   4659: 'Spare_Fault_4659', class No Acknowledgement, trigger "DB302_HMI_Faults_Carrier72_Faults_3" bit 2
   4660: 'Spare_Fault_4660', class No Acknowledgement, trigger "DB302_HMI_Faults_Carrier72_Faults_3" bit 3
   4661: 'Spare_Fault_4661', class No Acknowledgement, trigger "DB302_HMI_Faults_Carrier72_Faults_3" bit 4
   4662: 'Spare_Fault_4662', class No Acknowledgement, trigger "DB302_HMI_Faults_Carrier72_Faults_3" bit 5
   4663: 'Spare_Fault_4663', class No Acknowledgement, trigger "DB302_HMI_Faults_Carrier72_Faults_3" bit 6
   4664: 'Spare_Fault_4664', class No Acknowledgement, trigger "DB302_HMI_Faults_Carrier72_Faults_3" bit 7
   4665: 'Spare_Fault_4665', class No Acknowledgement, trigger "DB302_HMI_Faults_Carrier72_Faults_3" bit 8
   4666: 'Spare_Fault_4666', class No Acknowledgement, trigger "DB302_HMI_Faults_Carrier72_Faults_3" bit 9
   4667: 'Spare_Fault_4667', class No Acknowledgement, trigger "DB302_HMI_Faults_Carrier72_Faults_3" bit 10
   4668: 'Spare_Fault_4668', class No Acknowledgement, trigger "DB302_HMI_Faults_Carrier72_Faults_3" bit 11
   4669: 'Spare_Fault_4669', class No Acknowledgement, trigger "DB302_HMI_Faults_Carrier72_Faults_3" bit 12
   4670: 'Spare_Fault_4670', class No Acknowledgement, trigger "DB302_HMI_Faults_Carrier72_Faults_3" bit 13
   4671: 'Spare_Fault_4671', class No Acknowledgement, trigger "DB302_HMI_Faults_Carrier72_Faults_3" bit 14
   4672: 'Spare_Fault_4672', class No Acknowledgement, trigger "DB302_HMI_Faults_Carrier72_Faults_3" bit 15
   4673: 'Carrier 73 Disconnect Open Power Fault DI11.0', class No Acknowledgement, trigger "DB302_HMI_Faults_Carrier73_Faults_0" bit 0
   4674: 'Carrier 73 Drive Profinet Comm Fault', class No Acknowledgement, trigger "DB302_HMI_Faults_Carrier73_Faults_0" bit 1
   4675: 'Carrier 73 Production Stop Not Reset', class No Acknowledgement, trigger "DB302_HMI_Faults_Carrier73_Faults_0" bit 2
   4676: 'Carrier 73 CB02122 Tripped', class No Acknowledgement, trigger "DB302_HMI_Faults_Carrier73_Faults_0" bit 3
   4677: 'Carrier 73 CB02123 Tripped', class No Acknowledgement, trigger "DB302_HMI_Faults_Carrier73_Faults_0" bit 4
   4678: 'Carrier 73 AUX1 CB Tripped', class No Acknowledgement, trigger "DB302_HMI_Faults_Carrier73_Faults_0" bit 5
   4679: 'Carrier 73 AUX2 CB Tripped', class No Acknowledgement, trigger "DB302_HMI_Faults_Carrier73_Faults_0" bit 6
   4680: 'Carrier 73 PLC Not Communicating', class No Acknowledgement, trigger "DB302_HMI_Faults_Carrier73_Faults_0" bit 7
   4681: 'Carrier 73 Safe Input Card Fault', class No Acknowledgement, trigger "DB302_HMI_Faults_Carrier73_Faults_0" bit 8
   4682: 'Carrier 73 Safe Output Card Fault', class No Acknowledgement, trigger "DB302_HMI_Faults_Carrier73_Faults_0" bit 9
   4683: 'Carrier 73 Standard Input Card Fault', class No Acknowledgement, trigger "DB302_HMI_Faults_Carrier73_Faults_0" bit 10
   4684: 'Carrier 73 Standard Output Card Fault', class No Acknowledgement, trigger "DB302_HMI_Faults_Carrier73_Faults_0" bit 11
   4685: 'Carrier 73 Encoder Position Fault', class No Acknowledgement, trigger "DB302_HMI_Faults_Carrier73_Faults_0" bit 12
   4686: 'Carrier 73 Encoder Internal Error', class No Acknowledgement, trigger "DB302_HMI_Faults_Carrier73_Faults_0" bit 13
   4687: 'Carrier 73 Encoder Comm Fault', class No Acknowledgement, trigger "DB302_HMI_Faults_Carrier73_Faults_0" bit 14
   4688: 'Carrier 73 HMI Comm Fault', class No Acknowledgement, trigger "DB302_HMI_Faults_Carrier73_Faults_0" bit 15
   4689: 'Carrier 73 Crash Detection Fault', class No Acknowledgement, trigger "DB302_HMI_Faults_Carrier73_Faults_1" bit 0
   4690: 'Carrier 73 Carrier Number Invalid', class No Acknowledgement, trigger "DB302_HMI_Faults_Carrier73_Faults_1" bit 1
   4691: 'Carrier 73 Drive: PROFINET configuration error', class No Acknowledgement, trigger "DB302_HMI_Faults_Carrier73_Faults_1" bit 2
   4692: 'Carrier 73 Drive: Error internal communications', class No Acknowledgement, trigger "DB302_HMI_Faults_Carrier73_Faults_1" bit 3
   4693: 'Carrier 73 Drive: Motor overtemperature', class No Acknowledgement, trigger "DB302_HMI_Faults_Carrier73_Faults_1" bit 4
   4694: 'Carrier 73 Drive: Motor overcurrent', class No Acknowledgement, trigger "DB302_HMI_Faults_Carrier73_Faults_1" bit 5
   4695: 'Carrier 73 Drive: Infeed or power unit not ready', class No Acknowledgement, trigger "DB302_HMI_Faults_Carrier73_Faults_1" bit 6
   4696: 'Carrier 73 Drive: Short-circuit/ground fault detected', class No Acknowledgement, trigger "DB302_HMI_Faults_Carrier73_Faults_1" bit 7
   4697: 'Carrier 73 Drive: PROFINET Setpoint timeout', class No Acknowledgement, trigger "DB302_HMI_Faults_Carrier73_Faults_1" bit 8
   4698: 'Carrier 73 Power unit: Overcurrent', class No Acknowledgement, trigger "DB302_HMI_Faults_Carrier73_Faults_1" bit 9
   4699: 'Carrier 73 Power unit: DC link voltage overvoltage', class No Acknowledgement, trigger "DB302_HMI_Faults_Carrier73_Faults_1" bit 10
   4700: 'Carrier 73 Power unit: DC link voltage undervoltage', class No Acknowledgement, trigger "DB302_HMI_Faults_Carrier73_Faults_1" bit 11
   4701: 'Carrier 73 Power unit: Line phase failure in main circuit', class No Acknowledgement, trigger "DB302_HMI_Faults_Carrier73_Faults_1" bit 12
   4702: 'Carrier 73 Power unit: Phase failure motor cable', class No Acknowledgement, trigger "DB302_HMI_Faults_Carrier73_Faults_1" bit 13
   4703: 'Carrier 73 Power unit: Ground fault', class No Acknowledgement, trigger "DB302_HMI_Faults_Carrier73_Faults_1" bit 14
   4704: 'Spare_Fault_4704', class No Acknowledgement, trigger "DB302_HMI_Faults_Carrier73_Faults_1" bit 15
   4705: 'Carrier 73 Motion Off Fault', class No Acknowledgement, trigger "DB302_HMI_Faults_Carrier73_Faults_2" bit 0
   4706: 'Carrier 73 Motion On Fault', class No Acknowledgement, trigger "DB302_HMI_Faults_Carrier73_Faults_2" bit 1
   4707: 'Carrier 73 Spacing Fault', class No Acknowledgement, trigger "DB302_HMI_Faults_Carrier73_Faults_2" bit 2
   4708: 'Carrier 73 Duplicate Carrier Number Fault', class No Acknowledgement, trigger "DB302_HMI_Faults_Carrier73_Faults_2" bit 3
   4709: 'Spare_Fault_4709', class No Acknowledgement, trigger "DB302_HMI_Faults_Carrier73_Faults_2" bit 4
   4710: 'Spare_Fault_4710', class No Acknowledgement, trigger "DB302_HMI_Faults_Carrier73_Faults_2" bit 5
   4711: 'Spare_Fault_4711', class No Acknowledgement, trigger "DB302_HMI_Faults_Carrier73_Faults_2" bit 6
   4712: 'Spare_Fault_4712', class No Acknowledgement, trigger "DB302_HMI_Faults_Carrier73_Faults_2" bit 7
   4713: 'Spare_Fault_4713', class No Acknowledgement, trigger "DB302_HMI_Faults_Carrier73_Faults_2" bit 8
   4714: 'Spare_Fault_4714', class No Acknowledgement, trigger "DB302_HMI_Faults_Carrier73_Faults_2" bit 9
   4715: 'Spare_Fault_4715', class No Acknowledgement, trigger "DB302_HMI_Faults_Carrier73_Faults_2" bit 10
   4716: 'Spare_Fault_4716', class No Acknowledgement, trigger "DB302_HMI_Faults_Carrier73_Faults_2" bit 11
   4717: 'Spare_Fault_4717', class No Acknowledgement, trigger "DB302_HMI_Faults_Carrier73_Faults_2" bit 12
   4718: 'Spare_Fault_4718', class No Acknowledgement, trigger "DB302_HMI_Faults_Carrier73_Faults_2" bit 13
   4719: 'Spare_Fault_4719', class No Acknowledgement, trigger "DB302_HMI_Faults_Carrier73_Faults_2" bit 14
   4720: 'Spare_Fault_4720', class No Acknowledgement, trigger "DB302_HMI_Faults_Carrier73_Faults_2" bit 15
   4721: 'Spare_Fault_4721', class No Acknowledgement, trigger "DB302_HMI_Faults_Carrier73_Faults_3" bit 0
   4722: 'Spare_Fault_4722', class No Acknowledgement, trigger "DB302_HMI_Faults_Carrier73_Faults_3" bit 1
   4723: 'Spare_Fault_4723', class No Acknowledgement, trigger "DB302_HMI_Faults_Carrier73_Faults_3" bit 2
   4724: 'Spare_Fault_4724', class No Acknowledgement, trigger "DB302_HMI_Faults_Carrier73_Faults_3" bit 3
   4725: 'Spare_Fault_4725', class No Acknowledgement, trigger "DB302_HMI_Faults_Carrier73_Faults_3" bit 4
   4726: 'Spare_Fault_4726', class No Acknowledgement, trigger "DB302_HMI_Faults_Carrier73_Faults_3" bit 5
   4727: 'Spare_Fault_4727', class No Acknowledgement, trigger "DB302_HMI_Faults_Carrier73_Faults_3" bit 6
   4728: 'Spare_Fault_4728', class No Acknowledgement, trigger "DB302_HMI_Faults_Carrier73_Faults_3" bit 7
   4729: 'Spare_Fault_4729', class No Acknowledgement, trigger "DB302_HMI_Faults_Carrier73_Faults_3" bit 8
   4730: 'Spare_Fault_4730', class No Acknowledgement, trigger "DB302_HMI_Faults_Carrier73_Faults_3" bit 9
   4731: 'Spare_Fault_4731', class No Acknowledgement, trigger "DB302_HMI_Faults_Carrier73_Faults_3" bit 10
   4732: 'Spare_Fault_4732', class No Acknowledgement, trigger "DB302_HMI_Faults_Carrier73_Faults_3" bit 11
   4733: 'Spare_Fault_4733', class No Acknowledgement, trigger "DB302_HMI_Faults_Carrier73_Faults_3" bit 12
   4734: 'Spare_Fault_4734', class No Acknowledgement, trigger "DB302_HMI_Faults_Carrier73_Faults_3" bit 13
   4735: 'Spare_Fault_4735', class No Acknowledgement, trigger "DB302_HMI_Faults_Carrier73_Faults_3" bit 14
   4736: 'Spare_Fault_4736', class No Acknowledgement, trigger "DB302_HMI_Faults_Carrier73_Faults_3" bit 15
   4737: 'Carrier 74 Disconnect Open Power Fault DI11.0', class No Acknowledgement, trigger "DB302_HMI_Faults_Carrier74_Faults_0" bit 0
   4738: 'Carrier 74 Drive Profinet Comm Fault', class No Acknowledgement, trigger "DB302_HMI_Faults_Carrier74_Faults_0" bit 1
   4739: 'Carrier 74 Production Stop Not Reset', class No Acknowledgement, trigger "DB302_HMI_Faults_Carrier74_Faults_0" bit 2
   4740: 'Carrier 74 CB02122 Tripped', class No Acknowledgement, trigger "DB302_HMI_Faults_Carrier74_Faults_0" bit 3
   4741: 'Carrier 74 CB02123 Tripped', class No Acknowledgement, trigger "DB302_HMI_Faults_Carrier74_Faults_0" bit 4
   4742: 'Carrier 74 AUX1 CB Tripped', class No Acknowledgement, trigger "DB302_HMI_Faults_Carrier74_Faults_0" bit 5
   4743: 'Carrier 74 AUX2 CB Tripped', class No Acknowledgement, trigger "DB302_HMI_Faults_Carrier74_Faults_0" bit 6
   4744: 'Carrier 74 PLC Not Communicating', class No Acknowledgement, trigger "DB302_HMI_Faults_Carrier74_Faults_0" bit 7
   4745: 'Carrier 74 Safe Input Card Fault', class No Acknowledgement, trigger "DB302_HMI_Faults_Carrier74_Faults_0" bit 8
   4746: 'Carrier 74 Safe Output Card Fault', class No Acknowledgement, trigger "DB302_HMI_Faults_Carrier74_Faults_0" bit 9
   4747: 'Carrier 74 Standard Input Card Fault', class No Acknowledgement, trigger "DB302_HMI_Faults_Carrier74_Faults_0" bit 10
   4748: 'Carrier 74 Standard Output Card Fault', class No Acknowledgement, trigger "DB302_HMI_Faults_Carrier74_Faults_0" bit 11
   4749: 'Carrier 74 Encoder Position Fault', class No Acknowledgement, trigger "DB302_HMI_Faults_Carrier74_Faults_0" bit 12
   4750: 'Carrier 74 Encoder Internal Error', class No Acknowledgement, trigger "DB302_HMI_Faults_Carrier74_Faults_0" bit 13
   4751: 'Carrier 74 Encoder Comm Fault', class No Acknowledgement, trigger "DB302_HMI_Faults_Carrier74_Faults_0" bit 14
   4752: 'Carrier 74 HMI Comm Fault', class No Acknowledgement, trigger "DB302_HMI_Faults_Carrier74_Faults_0" bit 15
   4753: 'Carrier 74 Crash Detection Fault', class No Acknowledgement, trigger "DB302_HMI_Faults_Carrier74_Faults_1" bit 0
   4754: 'Carrier 74 Carrier Number Invalid', class No Acknowledgement, trigger "DB302_HMI_Faults_Carrier74_Faults_1" bit 1
   4755: 'Carrier 74 Drive: PROFINET configuration error', class No Acknowledgement, trigger "DB302_HMI_Faults_Carrier74_Faults_1" bit 2
   4756: 'Carrier 74 Drive: Error internal communications', class No Acknowledgement, trigger "DB302_HMI_Faults_Carrier74_Faults_1" bit 3
   4757: 'Carrier 74 Drive: Motor overtemperature', class No Acknowledgement, trigger "DB302_HMI_Faults_Carrier74_Faults_1" bit 4
   4758: 'Carrier 74 Drive: Motor overcurrent', class No Acknowledgement, trigger "DB302_HMI_Faults_Carrier74_Faults_1" bit 5
   4759: 'Carrier 74 Drive: Infeed or power unit not ready', class No Acknowledgement, trigger "DB302_HMI_Faults_Carrier74_Faults_1" bit 6
   4760: 'Carrier 74 Drive: Short-circuit/ground fault detected', class No Acknowledgement, trigger "DB302_HMI_Faults_Carrier74_Faults_1" bit 7
   4761: 'Carrier 74 Drive: PROFINET Setpoint timeout', class No Acknowledgement, trigger "DB302_HMI_Faults_Carrier74_Faults_1" bit 8
   4762: 'Carrier 74 Power unit: Overcurrent', class No Acknowledgement, trigger "DB302_HMI_Faults_Carrier74_Faults_1" bit 9
   4763: 'Carrier 74 Power unit: DC link voltage overvoltage', class No Acknowledgement, trigger "DB302_HMI_Faults_Carrier74_Faults_1" bit 10
   4764: 'Carrier 74 Power unit: DC link voltage undervoltage', class No Acknowledgement, trigger "DB302_HMI_Faults_Carrier74_Faults_1" bit 11
   4765: 'Carrier 74 Power unit: Line phase failure in main circuit', class No Acknowledgement, trigger "DB302_HMI_Faults_Carrier74_Faults_1" bit 12
   4766: 'Carrier 74 Power unit: Phase failure motor cable', class No Acknowledgement, trigger "DB302_HMI_Faults_Carrier74_Faults_1" bit 13
   4767: 'Carrier 74 Power unit: Ground fault', class No Acknowledgement, trigger "DB302_HMI_Faults_Carrier74_Faults_1" bit 14
   4768: 'Spare_Fault_4768', class No Acknowledgement, trigger "DB302_HMI_Faults_Carrier74_Faults_1" bit 15
   4769: 'Carrier 74 Motion Off Fault', class No Acknowledgement, trigger "DB302_HMI_Faults_Carrier74_Faults_2" bit 0
   4770: 'Carrier 74 Motion On Fault', class No Acknowledgement, trigger "DB302_HMI_Faults_Carrier74_Faults_2" bit 1
   4771: 'Carrier 74 Spacing Fault', class No Acknowledgement, trigger "DB302_HMI_Faults_Carrier74_Faults_2" bit 2
   4772: 'Carrier 74 Duplicate Carrier Number Fault', class No Acknowledgement, trigger "DB302_HMI_Faults_Carrier74_Faults_2" bit 3
   4773: 'Spare_Fault_4773', class No Acknowledgement, trigger "DB302_HMI_Faults_Carrier74_Faults_2" bit 4
   4774: 'Spare_Fault_4774', class No Acknowledgement, trigger "DB302_HMI_Faults_Carrier74_Faults_2" bit 5
   4775: 'Spare_Fault_4775', class No Acknowledgement, trigger "DB302_HMI_Faults_Carrier74_Faults_2" bit 6
   4776: 'Spare_Fault_4776', class No Acknowledgement, trigger "DB302_HMI_Faults_Carrier74_Faults_2" bit 7
   4777: 'Spare_Fault_4777', class No Acknowledgement, trigger "DB302_HMI_Faults_Carrier74_Faults_2" bit 8
   4778: 'Spare_Fault_4778', class No Acknowledgement, trigger "DB302_HMI_Faults_Carrier74_Faults_2" bit 9
   4779: 'Spare_Fault_4779', class No Acknowledgement, trigger "DB302_HMI_Faults_Carrier74_Faults_2" bit 10
   4780: 'Spare_Fault_4780', class No Acknowledgement, trigger "DB302_HMI_Faults_Carrier74_Faults_2" bit 11
   4781: 'Spare_Fault_4781', class No Acknowledgement, trigger "DB302_HMI_Faults_Carrier74_Faults_2" bit 12
   4782: 'Spare_Fault_4782', class No Acknowledgement, trigger "DB302_HMI_Faults_Carrier74_Faults_2" bit 13
   4783: 'Spare_Fault_4783', class No Acknowledgement, trigger "DB302_HMI_Faults_Carrier74_Faults_2" bit 14
   4784: 'Spare_Fault_4784', class No Acknowledgement, trigger "DB302_HMI_Faults_Carrier74_Faults_2" bit 15
   4785: 'Spare_Fault_4785', class No Acknowledgement, trigger "DB302_HMI_Faults_Carrier74_Faults_3" bit 0
   4786: 'Spare_Fault_4786', class No Acknowledgement, trigger "DB302_HMI_Faults_Carrier74_Faults_3" bit 1
   4787: 'Spare_Fault_4787', class No Acknowledgement, trigger "DB302_HMI_Faults_Carrier74_Faults_3" bit 2
   4788: 'Spare_Fault_4788', class No Acknowledgement, trigger "DB302_HMI_Faults_Carrier74_Faults_3" bit 3
   4789: 'Spare_Fault_4789', class No Acknowledgement, trigger "DB302_HMI_Faults_Carrier74_Faults_3" bit 4
   4790: 'Spare_Fault_4790', class No Acknowledgement, trigger "DB302_HMI_Faults_Carrier74_Faults_3" bit 5
   4791: 'Spare_Fault_4791', class No Acknowledgement, trigger "DB302_HMI_Faults_Carrier74_Faults_3" bit 6
   4792: 'Spare_Fault_4792', class No Acknowledgement, trigger "DB302_HMI_Faults_Carrier74_Faults_3" bit 7
   4793: 'Spare_Fault_4793', class No Acknowledgement, trigger "DB302_HMI_Faults_Carrier74_Faults_3" bit 8
   4794: 'Spare_Fault_4794', class No Acknowledgement, trigger "DB302_HMI_Faults_Carrier74_Faults_3" bit 9
   4795: 'Spare_Fault_4795', class No Acknowledgement, trigger "DB302_HMI_Faults_Carrier74_Faults_3" bit 10
   4796: 'Spare_Fault_4796', class No Acknowledgement, trigger "DB302_HMI_Faults_Carrier74_Faults_3" bit 11
   4797: 'Spare_Fault_4797', class No Acknowledgement, trigger "DB302_HMI_Faults_Carrier74_Faults_3" bit 12
   4798: 'Spare_Fault_4798', class No Acknowledgement, trigger "DB302_HMI_Faults_Carrier74_Faults_3" bit 13
   4799: 'Spare_Fault_4799', class No Acknowledgement, trigger "DB302_HMI_Faults_Carrier74_Faults_3" bit 14
   4800: 'Spare_Fault_4800', class No Acknowledgement, trigger "DB302_HMI_Faults_Carrier74_Faults_3" bit 15
   4801: 'Carrier 75 Disconnect Open Power Fault DI11.0', class No Acknowledgement, trigger "DB302_HMI_Faults_Carrier75_Faults_0" bit 0
   4802: 'Carrier 75 Drive Profinet Comm Fault', class No Acknowledgement, trigger "DB302_HMI_Faults_Carrier75_Faults_0" bit 1
   4803: 'Carrier 75 Production Stop Not Reset', class No Acknowledgement, trigger "DB302_HMI_Faults_Carrier75_Faults_0" bit 2
   4804: 'Carrier 75 CB02122 Tripped', class No Acknowledgement, trigger "DB302_HMI_Faults_Carrier75_Faults_0" bit 3
   4805: 'Carrier 75 CB02123 Tripped', class No Acknowledgement, trigger "DB302_HMI_Faults_Carrier75_Faults_0" bit 4
   4806: 'Carrier 75 AUX1 CB Tripped', class No Acknowledgement, trigger "DB302_HMI_Faults_Carrier75_Faults_0" bit 5
   4807: 'Carrier 75 AUX2 CB Tripped', class No Acknowledgement, trigger "DB302_HMI_Faults_Carrier75_Faults_0" bit 6
   4808: 'Carrier 75 PLC Not Communicating', class No Acknowledgement, trigger "DB302_HMI_Faults_Carrier75_Faults_0" bit 7
   4809: 'Carrier 75 Safe Input Card Fault', class No Acknowledgement, trigger "DB302_HMI_Faults_Carrier75_Faults_0" bit 8
   4810: 'Carrier 75 Safe Output Card Fault', class No Acknowledgement, trigger "DB302_HMI_Faults_Carrier75_Faults_0" bit 9
   4811: 'Carrier 75 Standard Input Card Fault', class No Acknowledgement, trigger "DB302_HMI_Faults_Carrier75_Faults_0" bit 10
   4812: 'Carrier 75 Standard Output Card Fault', class No Acknowledgement, trigger "DB302_HMI_Faults_Carrier75_Faults_0" bit 11
   4813: 'Carrier 75 Encoder Position Fault', class No Acknowledgement, trigger "DB302_HMI_Faults_Carrier75_Faults_0" bit 12
   4814: 'Carrier 75 Encoder Internal Error', class No Acknowledgement, trigger "DB302_HMI_Faults_Carrier75_Faults_0" bit 13
   4815: 'Carrier 75 Encoder Comm Fault', class No Acknowledgement, trigger "DB302_HMI_Faults_Carrier75_Faults_0" bit 14
   4816: 'Carrier 75 HMI Comm Fault', class No Acknowledgement, trigger "DB302_HMI_Faults_Carrier75_Faults_0" bit 15
   4817: 'Carrier 75 Crash Detection Fault', class No Acknowledgement, trigger "DB302_HMI_Faults_Carrier75_Faults_1" bit 0
   4818: 'Carrier 75 Carrier Number Invalid', class No Acknowledgement, trigger "DB302_HMI_Faults_Carrier75_Faults_1" bit 1
   4819: 'Carrier 75 Drive: PROFINET configuration error', class No Acknowledgement, trigger "DB302_HMI_Faults_Carrier75_Faults_1" bit 2
   4820: 'Carrier 75 Drive: Error internal communications', class No Acknowledgement, trigger "DB302_HMI_Faults_Carrier75_Faults_1" bit 3
   4821: 'Carrier 75 Drive: Motor overtemperature', class No Acknowledgement, trigger "DB302_HMI_Faults_Carrier75_Faults_1" bit 4
   4822: 'Carrier 75 Drive: Motor overcurrent', class No Acknowledgement, trigger "DB302_HMI_Faults_Carrier75_Faults_1" bit 5
   4823: 'Carrier 75 Drive: Infeed or power unit not ready', class No Acknowledgement, trigger "DB302_HMI_Faults_Carrier75_Faults_1" bit 6
   4824: 'Carrier 75 Drive: Short-circuit/ground fault detected', class No Acknowledgement, trigger "DB302_HMI_Faults_Carrier75_Faults_1" bit 7
   4825: 'Carrier 75 Drive: PROFINET Setpoint timeout', class No Acknowledgement, trigger "DB302_HMI_Faults_Carrier75_Faults_1" bit 8
   4826: 'Carrier 75 Power unit: Overcurrent', class No Acknowledgement, trigger "DB302_HMI_Faults_Carrier75_Faults_1" bit 9
   4827: 'Carrier 75 Power unit: DC link voltage overvoltage', class No Acknowledgement, trigger "DB302_HMI_Faults_Carrier75_Faults_1" bit 10
   4828: 'Carrier 75 Power unit: DC link voltage undervoltage', class No Acknowledgement, trigger "DB302_HMI_Faults_Carrier75_Faults_1" bit 11
   4829: 'Carrier 75 Power unit: Line phase failure in main circuit', class No Acknowledgement, trigger "DB302_HMI_Faults_Carrier75_Faults_1" bit 12
   4830: 'Carrier 75 Power unit: Phase failure motor cable', class No Acknowledgement, trigger "DB302_HMI_Faults_Carrier75_Faults_1" bit 13
   4831: 'Carrier 75 Power unit: Ground fault', class No Acknowledgement, trigger "DB302_HMI_Faults_Carrier75_Faults_1" bit 14
   4832: 'Spare_Fault_4832', class No Acknowledgement, trigger "DB302_HMI_Faults_Carrier75_Faults_1" bit 15
   4833: 'Carrier 75 Motion Off Fault', class No Acknowledgement, trigger "DB302_HMI_Faults_Carrier75_Faults_2" bit 0
   4834: 'Carrier 75 Motion On Fault', class No Acknowledgement, trigger "DB302_HMI_Faults_Carrier75_Faults_2" bit 1
   4835: 'Carrier 75 Spacing Fault', class No Acknowledgement, trigger "DB302_HMI_Faults_Carrier75_Faults_2" bit 2
   4836: 'Carrier 75 Duplicate Carrier Number Fault', class No Acknowledgement, trigger "DB302_HMI_Faults_Carrier75_Faults_2" bit 3
   4837: 'Spare_Fault_4837', class No Acknowledgement, trigger "DB302_HMI_Faults_Carrier75_Faults_2" bit 4
   4838: 'Spare_Fault_4838', class No Acknowledgement, trigger "DB302_HMI_Faults_Carrier75_Faults_2" bit 5
   4839: 'Spare_Fault_4839', class No Acknowledgement, trigger "DB302_HMI_Faults_Carrier75_Faults_2" bit 6
   4840: 'Spare_Fault_4840', class No Acknowledgement, trigger "DB302_HMI_Faults_Carrier75_Faults_2" bit 7
   4841: 'Spare_Fault_4841', class No Acknowledgement, trigger "DB302_HMI_Faults_Carrier75_Faults_2" bit 8
   4842: 'Spare_Fault_4842', class No Acknowledgement, trigger "DB302_HMI_Faults_Carrier75_Faults_2" bit 9
   4843: 'Spare_Fault_4843', class No Acknowledgement, trigger "DB302_HMI_Faults_Carrier75_Faults_2" bit 10
   4844: 'Spare_Fault_4844', class No Acknowledgement, trigger "DB302_HMI_Faults_Carrier75_Faults_2" bit 11
   4845: 'Spare_Fault_4845', class No Acknowledgement, trigger "DB302_HMI_Faults_Carrier75_Faults_2" bit 12
   4846: 'Spare_Fault_4846', class No Acknowledgement, trigger "DB302_HMI_Faults_Carrier75_Faults_2" bit 13
   4847: 'Spare_Fault_4847', class No Acknowledgement, trigger "DB302_HMI_Faults_Carrier75_Faults_2" bit 14
   4848: 'Spare_Fault_4848', class No Acknowledgement, trigger "DB302_HMI_Faults_Carrier75_Faults_2" bit 15
   4849: 'Spare_Fault_4849', class No Acknowledgement, trigger "DB302_HMI_Faults_Carrier75_Faults_3" bit 0
   4850: 'Spare_Fault_4850', class No Acknowledgement, trigger "DB302_HMI_Faults_Carrier75_Faults_3" bit 1
   4851: 'Spare_Fault_4851', class No Acknowledgement, trigger "DB302_HMI_Faults_Carrier75_Faults_3" bit 2
   4852: 'Spare_Fault_4852', class No Acknowledgement, trigger "DB302_HMI_Faults_Carrier75_Faults_3" bit 3
   4853: 'Spare_Fault_4853', class No Acknowledgement, trigger "DB302_HMI_Faults_Carrier75_Faults_3" bit 4
   4854: 'Spare_Fault_4854', class No Acknowledgement, trigger "DB302_HMI_Faults_Carrier75_Faults_3" bit 5
   4855: 'Spare_Fault_4855', class No Acknowledgement, trigger "DB302_HMI_Faults_Carrier75_Faults_3" bit 6
   4856: 'Spare_Fault_4856', class No Acknowledgement, trigger "DB302_HMI_Faults_Carrier75_Faults_3" bit 7
   4857: 'Spare_Fault_4857', class No Acknowledgement, trigger "DB302_HMI_Faults_Carrier75_Faults_3" bit 8
   4858: 'Spare_Fault_4858', class No Acknowledgement, trigger "DB302_HMI_Faults_Carrier75_Faults_3" bit 9
   4859: 'Spare_Fault_4859', class No Acknowledgement, trigger "DB302_HMI_Faults_Carrier75_Faults_3" bit 10
   4860: 'Spare_Fault_4860', class No Acknowledgement, trigger "DB302_HMI_Faults_Carrier75_Faults_3" bit 11
   4861: 'Spare_Fault_4861', class No Acknowledgement, trigger "DB302_HMI_Faults_Carrier75_Faults_3" bit 12
   4862: 'Spare_Fault_4862', class No Acknowledgement, trigger "DB302_HMI_Faults_Carrier75_Faults_3" bit 13
   4863: 'Spare_Fault_4863', class No Acknowledgement, trigger "DB302_HMI_Faults_Carrier75_Faults_3" bit 14
   4864: 'Spare_Fault_4864', class No Acknowledgement, trigger "DB302_HMI_Faults_Carrier75_Faults_3" bit 15
   4865: 'Carrier 76 Disconnect Open Power Fault DI11.0', class No Acknowledgement, trigger "DB302_HMI_Faults_Carrier76_Faults_0" bit 0
   4866: 'Carrier 76 Drive Profinet Comm Fault', class No Acknowledgement, trigger "DB302_HMI_Faults_Carrier76_Faults_0" bit 1
   4867: 'Carrier 76 Production Stop Not Reset', class No Acknowledgement, trigger "DB302_HMI_Faults_Carrier76_Faults_0" bit 2
   4868: 'Carrier 76 CB02122 Tripped', class No Acknowledgement, trigger "DB302_HMI_Faults_Carrier76_Faults_0" bit 3
   4869: 'Carrier 76 CB02123 Tripped', class No Acknowledgement, trigger "DB302_HMI_Faults_Carrier76_Faults_0" bit 4
   4870: 'Carrier 76 AUX1 CB Tripped', class No Acknowledgement, trigger "DB302_HMI_Faults_Carrier76_Faults_0" bit 5
   4871: 'Carrier 76 AUX2 CB Tripped', class No Acknowledgement, trigger "DB302_HMI_Faults_Carrier76_Faults_0" bit 6
   4872: 'Carrier 76 PLC Not Communicating', class No Acknowledgement, trigger "DB302_HMI_Faults_Carrier76_Faults_0" bit 7
   4873: 'Carrier 76 Safe Input Card Fault', class No Acknowledgement, trigger "DB302_HMI_Faults_Carrier76_Faults_0" bit 8
   4874: 'Carrier 76 Safe Output Card Fault', class No Acknowledgement, trigger "DB302_HMI_Faults_Carrier76_Faults_0" bit 9
   4875: 'Carrier 76 Standard Input Card Fault', class No Acknowledgement, trigger "DB302_HMI_Faults_Carrier76_Faults_0" bit 10
   4876: 'Carrier 76 Standard Output Card Fault', class No Acknowledgement, trigger "DB302_HMI_Faults_Carrier76_Faults_0" bit 11
   4877: 'Carrier 76 Encoder Position Fault', class No Acknowledgement, trigger "DB302_HMI_Faults_Carrier76_Faults_0" bit 12
   4878: 'Carrier 76 Encoder Internal Error', class No Acknowledgement, trigger "DB302_HMI_Faults_Carrier76_Faults_0" bit 13
   4879: 'Carrier 76 Encoder Comm Fault', class No Acknowledgement, trigger "DB302_HMI_Faults_Carrier76_Faults_0" bit 14
   4880: 'Carrier 76 HMI Comm Fault', class No Acknowledgement, trigger "DB302_HMI_Faults_Carrier76_Faults_0" bit 15
   4881: 'Carrier 76 Crash Detection Fault', class No Acknowledgement, trigger "DB302_HMI_Faults_Carrier76_Faults_1" bit 0
   4882: 'Carrier 76 Carrier Number Invalid', class No Acknowledgement, trigger "DB302_HMI_Faults_Carrier76_Faults_1" bit 1
   4883: 'Carrier 76 Drive: PROFINET configuration error', class No Acknowledgement, trigger "DB302_HMI_Faults_Carrier76_Faults_1" bit 2
   4884: 'Carrier 76 Drive: Error internal communications', class No Acknowledgement, trigger "DB302_HMI_Faults_Carrier76_Faults_1" bit 3
   4885: 'Carrier 76 Drive: Motor overtemperature', class No Acknowledgement, trigger "DB302_HMI_Faults_Carrier76_Faults_1" bit 4
   4886: 'Carrier 76 Drive: Motor overcurrent', class No Acknowledgement, trigger "DB302_HMI_Faults_Carrier76_Faults_1" bit 5
   4887: 'Carrier 76 Drive: Infeed or power unit not ready', class No Acknowledgement, trigger "DB302_HMI_Faults_Carrier76_Faults_1" bit 6
   4888: 'Carrier 76 Drive: Short-circuit/ground fault detected', class No Acknowledgement, trigger "DB302_HMI_Faults_Carrier76_Faults_1" bit 7
   4889: 'Carrier 76 Drive: PROFINET Setpoint timeout', class No Acknowledgement, trigger "DB302_HMI_Faults_Carrier76_Faults_1" bit 8
   4890: 'Carrier 76 Power unit: Overcurrent', class No Acknowledgement, trigger "DB302_HMI_Faults_Carrier76_Faults_1" bit 9
   4891: 'Carrier 76 Power unit: DC link voltage overvoltage', class No Acknowledgement, trigger "DB302_HMI_Faults_Carrier76_Faults_1" bit 10
   4892: 'Carrier 76 Power unit: DC link voltage undervoltage', class No Acknowledgement, trigger "DB302_HMI_Faults_Carrier76_Faults_1" bit 11
   4893: 'Carrier 76 Power unit: Line phase failure in main circuit', class No Acknowledgement, trigger "DB302_HMI_Faults_Carrier76_Faults_1" bit 12
   4894: 'Carrier 76 Power unit: Phase failure motor cable', class No Acknowledgement, trigger "DB302_HMI_Faults_Carrier76_Faults_1" bit 13
   4895: 'Carrier 76 Power unit: Ground fault', class No Acknowledgement, trigger "DB302_HMI_Faults_Carrier76_Faults_1" bit 14
   4896: 'Spare_Fault_4896', class No Acknowledgement, trigger "DB302_HMI_Faults_Carrier76_Faults_1" bit 15
   4897: 'Carrier 76 Motion Off Fault', class No Acknowledgement, trigger "DB302_HMI_Faults_Carrier76_Faults_2" bit 0
   4898: 'Carrier 76 Motion On Fault', class No Acknowledgement, trigger "DB302_HMI_Faults_Carrier76_Faults_2" bit 1
   4899: 'Carrier 76 Spacing Fault', class No Acknowledgement, trigger "DB302_HMI_Faults_Carrier76_Faults_2" bit 2
   4900: 'Carrier 76 Duplicate Carrier Number Fault', class No Acknowledgement, trigger "DB302_HMI_Faults_Carrier76_Faults_2" bit 3
   4901: 'Spare_Fault_4901', class No Acknowledgement, trigger "DB302_HMI_Faults_Carrier76_Faults_2" bit 4
   4902: 'Spare_Fault_4902', class No Acknowledgement, trigger "DB302_HMI_Faults_Carrier76_Faults_2" bit 5
   4903: 'Spare_Fault_4903', class No Acknowledgement, trigger "DB302_HMI_Faults_Carrier76_Faults_2" bit 6
   4904: 'Spare_Fault_4904', class No Acknowledgement, trigger "DB302_HMI_Faults_Carrier76_Faults_2" bit 7
   4905: 'Spare_Fault_4905', class No Acknowledgement, trigger "DB302_HMI_Faults_Carrier76_Faults_2" bit 8
   4906: 'Spare_Fault_4906', class No Acknowledgement, trigger "DB302_HMI_Faults_Carrier76_Faults_2" bit 9
   4907: 'Spare_Fault_4907', class No Acknowledgement, trigger "DB302_HMI_Faults_Carrier76_Faults_2" bit 10
   4908: 'Spare_Fault_4908', class No Acknowledgement, trigger "DB302_HMI_Faults_Carrier76_Faults_2" bit 11
   4909: 'Spare_Fault_4909', class No Acknowledgement, trigger "DB302_HMI_Faults_Carrier76_Faults_2" bit 12
   4910: 'Spare_Fault_4910', class No Acknowledgement, trigger "DB302_HMI_Faults_Carrier76_Faults_2" bit 13
   4911: 'Spare_Fault_4911', class No Acknowledgement, trigger "DB302_HMI_Faults_Carrier76_Faults_2" bit 14
   4912: 'Spare_Fault_4912', class No Acknowledgement, trigger "DB302_HMI_Faults_Carrier76_Faults_2" bit 15
   4913: 'Spare_Fault_4913', class No Acknowledgement, trigger "DB302_HMI_Faults_Carrier76_Faults_3" bit 0
   4914: 'Spare_Fault_4914', class No Acknowledgement, trigger "DB302_HMI_Faults_Carrier76_Faults_3" bit 1
   4915: 'Spare_Fault_4915', class No Acknowledgement, trigger "DB302_HMI_Faults_Carrier76_Faults_3" bit 2
   4916: 'Spare_Fault_4916', class No Acknowledgement, trigger "DB302_HMI_Faults_Carrier76_Faults_3" bit 3
   4917: 'Spare_Fault_4917', class No Acknowledgement, trigger "DB302_HMI_Faults_Carrier76_Faults_3" bit 4
   4918: 'Spare_Fault_4918', class No Acknowledgement, trigger "DB302_HMI_Faults_Carrier76_Faults_3" bit 5
   4919: 'Spare_Fault_4919', class No Acknowledgement, trigger "DB302_HMI_Faults_Carrier76_Faults_3" bit 6
   4920: 'Spare_Fault_4920', class No Acknowledgement, trigger "DB302_HMI_Faults_Carrier76_Faults_3" bit 7
   4921: 'Spare_Fault_4921', class No Acknowledgement, trigger "DB302_HMI_Faults_Carrier76_Faults_3" bit 8
   4922: 'Spare_Fault_4922', class No Acknowledgement, trigger "DB302_HMI_Faults_Carrier76_Faults_3" bit 9
   4923: 'Spare_Fault_4923', class No Acknowledgement, trigger "DB302_HMI_Faults_Carrier76_Faults_3" bit 10
   4924: 'Spare_Fault_4924', class No Acknowledgement, trigger "DB302_HMI_Faults_Carrier76_Faults_3" bit 11
   4925: 'Spare_Fault_4925', class No Acknowledgement, trigger "DB302_HMI_Faults_Carrier76_Faults_3" bit 12
   4926: 'Spare_Fault_4926', class No Acknowledgement, trigger "DB302_HMI_Faults_Carrier76_Faults_3" bit 13
   4927: 'Spare_Fault_4927', class No Acknowledgement, trigger "DB302_HMI_Faults_Carrier76_Faults_3" bit 14
   4928: 'Spare_Fault_4928', class No Acknowledgement, trigger "DB302_HMI_Faults_Carrier76_Faults_3" bit 15
   4929: 'Carrier 77 Disconnect Open Power Fault DI11.0', class No Acknowledgement, trigger "DB302_HMI_Faults_Carrier77_Faults_0" bit 0
   4930: 'Carrier 77 Drive Profinet Comm Fault', class No Acknowledgement, trigger "DB302_HMI_Faults_Carrier77_Faults_0" bit 1
   4931: 'Carrier 77 Production Stop Not Reset', class No Acknowledgement, trigger "DB302_HMI_Faults_Carrier77_Faults_0" bit 2
   4932: 'Carrier 77 CB02122 Tripped', class No Acknowledgement, trigger "DB302_HMI_Faults_Carrier77_Faults_0" bit 3
   4933: 'Carrier 77 CB02123 Tripped', class No Acknowledgement, trigger "DB302_HMI_Faults_Carrier77_Faults_0" bit 4
   4934: 'Carrier 77 AUX1 CB Tripped', class No Acknowledgement, trigger "DB302_HMI_Faults_Carrier77_Faults_0" bit 5
   4935: 'Carrier 77 AUX2 CB Tripped', class No Acknowledgement, trigger "DB302_HMI_Faults_Carrier77_Faults_0" bit 6
   4936: 'Carrier 77 PLC Not Communicating', class No Acknowledgement, trigger "DB302_HMI_Faults_Carrier77_Faults_0" bit 7
   4937: 'Carrier 77 Safe Input Card Fault', class No Acknowledgement, trigger "DB302_HMI_Faults_Carrier77_Faults_0" bit 8
   4938: 'Carrier 77 Safe Output Card Fault', class No Acknowledgement, trigger "DB302_HMI_Faults_Carrier77_Faults_0" bit 9
   4939: 'Carrier 77 Standard Input Card Fault', class No Acknowledgement, trigger "DB302_HMI_Faults_Carrier77_Faults_0" bit 10
   4940: 'Carrier 77 Standard Output Card Fault', class No Acknowledgement, trigger "DB302_HMI_Faults_Carrier77_Faults_0" bit 11
   4941: 'Carrier 77 Encoder Position Fault', class No Acknowledgement, trigger "DB302_HMI_Faults_Carrier77_Faults_0" bit 12
   4942: 'Carrier 77 Encoder Internal Error', class No Acknowledgement, trigger "DB302_HMI_Faults_Carrier77_Faults_0" bit 13
   4943: 'Carrier 77 Encoder Comm Fault', class No Acknowledgement, trigger "DB302_HMI_Faults_Carrier77_Faults_0" bit 14
   4944: 'Carrier 77 HMI Comm Fault', class No Acknowledgement, trigger "DB302_HMI_Faults_Carrier77_Faults_0" bit 15
   4945: 'Carrier 77 Crash Detection Fault', class No Acknowledgement, trigger "DB302_HMI_Faults_Carrier77_Faults_1" bit 0
   4946: 'Carrier 77 Carrier Number Invalid', class No Acknowledgement, trigger "DB302_HMI_Faults_Carrier77_Faults_1" bit 1
   4947: 'Carrier 77 Drive: PROFINET configuration error', class No Acknowledgement, trigger "DB302_HMI_Faults_Carrier77_Faults_1" bit 2
   4948: 'Carrier 77 Drive: Error internal communications', class No Acknowledgement, trigger "DB302_HMI_Faults_Carrier77_Faults_1" bit 3
   4949: 'Carrier 77 Drive: Motor overtemperature', class No Acknowledgement, trigger "DB302_HMI_Faults_Carrier77_Faults_1" bit 4
   4950: 'Carrier 77 Drive: Motor overcurrent', class No Acknowledgement, trigger "DB302_HMI_Faults_Carrier77_Faults_1" bit 5
   4951: 'Carrier 77 Drive: Infeed or power unit not ready', class No Acknowledgement, trigger "DB302_HMI_Faults_Carrier77_Faults_1" bit 6
   4952: 'Carrier 77 Drive: Short-circuit/ground fault detected', class No Acknowledgement, trigger "DB302_HMI_Faults_Carrier77_Faults_1" bit 7
   4953: 'Carrier 77 Drive: PROFINET Setpoint timeout', class No Acknowledgement, trigger "DB302_HMI_Faults_Carrier77_Faults_1" bit 8
   4954: 'Carrier 77 Power unit: Overcurrent', class No Acknowledgement, trigger "DB302_HMI_Faults_Carrier77_Faults_1" bit 9
   4955: 'Carrier 77 Power unit: DC link voltage overvoltage', class No Acknowledgement, trigger "DB302_HMI_Faults_Carrier77_Faults_1" bit 10
   4956: 'Carrier 77 Power unit: DC link voltage undervoltage', class No Acknowledgement, trigger "DB302_HMI_Faults_Carrier77_Faults_1" bit 11
   4957: 'Carrier 77 Power unit: Line phase failure in main circuit', class No Acknowledgement, trigger "DB302_HMI_Faults_Carrier77_Faults_1" bit 12
   4958: 'Carrier 77 Power unit: Phase failure motor cable', class No Acknowledgement, trigger "DB302_HMI_Faults_Carrier77_Faults_1" bit 13
   4959: 'Carrier 77 Power unit: Ground fault', class No Acknowledgement, trigger "DB302_HMI_Faults_Carrier77_Faults_1" bit 14
   4960: 'Spare_Fault_4960', class No Acknowledgement, trigger "DB302_HMI_Faults_Carrier77_Faults_1" bit 15
   4961: 'Carrier 77 Motion Off Fault', class No Acknowledgement, trigger "DB302_HMI_Faults_Carrier77_Faults_2" bit 0
   4962: 'Carrier 77 Motion On Fault', class No Acknowledgement, trigger "DB302_HMI_Faults_Carrier77_Faults_2" bit 1
   4963: 'Carrier 77 Spacing Fault', class No Acknowledgement, trigger "DB302_HMI_Faults_Carrier77_Faults_2" bit 2
   4964: 'Carrier 77 Duplicate Carrier Number Fault', class No Acknowledgement, trigger "DB302_HMI_Faults_Carrier77_Faults_2" bit 3
   4965: 'Spare_Fault_4965', class No Acknowledgement, trigger "DB302_HMI_Faults_Carrier77_Faults_2" bit 4
   4966: 'Spare_Fault_4966', class No Acknowledgement, trigger "DB302_HMI_Faults_Carrier77_Faults_2" bit 5
   4967: 'Spare_Fault_4967', class No Acknowledgement, trigger "DB302_HMI_Faults_Carrier77_Faults_2" bit 6
   4968: 'Spare_Fault_4968', class No Acknowledgement, trigger "DB302_HMI_Faults_Carrier77_Faults_2" bit 7
   4969: 'Spare_Fault_4969', class No Acknowledgement, trigger "DB302_HMI_Faults_Carrier77_Faults_2" bit 8
   4970: 'Spare_Fault_4970', class No Acknowledgement, trigger "DB302_HMI_Faults_Carrier77_Faults_2" bit 9
   4971: 'Spare_Fault_4971', class No Acknowledgement, trigger "DB302_HMI_Faults_Carrier77_Faults_2" bit 10
   4972: 'Spare_Fault_4972', class No Acknowledgement, trigger "DB302_HMI_Faults_Carrier77_Faults_2" bit 11
   4973: 'Spare_Fault_4973', class No Acknowledgement, trigger "DB302_HMI_Faults_Carrier77_Faults_2" bit 12
   4974: 'Spare_Fault_4974', class No Acknowledgement, trigger "DB302_HMI_Faults_Carrier77_Faults_2" bit 13
   4975: 'Spare_Fault_4975', class No Acknowledgement, trigger "DB302_HMI_Faults_Carrier77_Faults_2" bit 14
   4976: 'Spare_Fault_4976', class No Acknowledgement, trigger "DB302_HMI_Faults_Carrier77_Faults_2" bit 15
   4977: 'Spare_Fault_4977', class No Acknowledgement, trigger "DB302_HMI_Faults_Carrier77_Faults_3" bit 0
   4978: 'Spare_Fault_4978', class No Acknowledgement, trigger "DB302_HMI_Faults_Carrier77_Faults_3" bit 1
   4979: 'Spare_Fault_4979', class No Acknowledgement, trigger "DB302_HMI_Faults_Carrier77_Faults_3" bit 2
   4980: 'Spare_Fault_4980', class No Acknowledgement, trigger "DB302_HMI_Faults_Carrier77_Faults_3" bit 3
   4981: 'Spare_Fault_4981', class No Acknowledgement, trigger "DB302_HMI_Faults_Carrier77_Faults_3" bit 4
   4982: 'Spare_Fault_4982', class No Acknowledgement, trigger "DB302_HMI_Faults_Carrier77_Faults_3" bit 5
   4983: 'Spare_Fault_4983', class No Acknowledgement, trigger "DB302_HMI_Faults_Carrier77_Faults_3" bit 6
   4984: 'Spare_Fault_4984', class No Acknowledgement, trigger "DB302_HMI_Faults_Carrier77_Faults_3" bit 7
   4985: 'Spare_Fault_4985', class No Acknowledgement, trigger "DB302_HMI_Faults_Carrier77_Faults_3" bit 8
   4986: 'Spare_Fault_4986', class No Acknowledgement, trigger "DB302_HMI_Faults_Carrier77_Faults_3" bit 9
   4987: 'Spare_Fault_4987', class No Acknowledgement, trigger "DB302_HMI_Faults_Carrier77_Faults_3" bit 10
   4988: 'Spare_Fault_4988', class No Acknowledgement, trigger "DB302_HMI_Faults_Carrier77_Faults_3" bit 11
   4989: 'Spare_Fault_4989', class No Acknowledgement, trigger "DB302_HMI_Faults_Carrier77_Faults_3" bit 12
   4990: 'Spare_Fault_4990', class No Acknowledgement, trigger "DB302_HMI_Faults_Carrier77_Faults_3" bit 13
   4991: 'Spare_Fault_4991', class No Acknowledgement, trigger "DB302_HMI_Faults_Carrier77_Faults_3" bit 14
   4992: 'Spare_Fault_4992', class No Acknowledgement, trigger "DB302_HMI_Faults_Carrier77_Faults_3" bit 15
   4993: 'Carrier 78 Disconnect Open Power Fault DI11.0', class No Acknowledgement, trigger "DB302_HMI_Faults_Carrier78_Faults_0" bit 0
   4994: 'Carrier 78 Drive Profinet Comm Fault', class No Acknowledgement, trigger "DB302_HMI_Faults_Carrier78_Faults_0" bit 1
   4995: 'Carrier 78 Production Stop Not Reset', class No Acknowledgement, trigger "DB302_HMI_Faults_Carrier78_Faults_0" bit 2
   4996: 'Carrier 78 CB02122 Tripped', class No Acknowledgement, trigger "DB302_HMI_Faults_Carrier78_Faults_0" bit 3
   4997: 'Carrier 78 CB02123 Tripped', class No Acknowledgement, trigger "DB302_HMI_Faults_Carrier78_Faults_0" bit 4
   4998: 'Carrier 78 AUX1 CB Tripped', class No Acknowledgement, trigger "DB302_HMI_Faults_Carrier78_Faults_0" bit 5
   4999: 'Carrier 78 AUX2 CB Tripped', class No Acknowledgement, trigger "DB302_HMI_Faults_Carrier78_Faults_0" bit 6
   5000: 'Carrier 78 PLC Not Communicating', class No Acknowledgement, trigger "DB302_HMI_Faults_Carrier78_Faults_0" bit 7
   5001: 'Carrier 78 Safe Input Card Fault', class No Acknowledgement, trigger "DB302_HMI_Faults_Carrier78_Faults_0" bit 8
   5002: 'Carrier 78 Safe Output Card Fault', class No Acknowledgement, trigger "DB302_HMI_Faults_Carrier78_Faults_0" bit 9
   5003: 'Carrier 78 Standard Input Card Fault', class No Acknowledgement, trigger "DB302_HMI_Faults_Carrier78_Faults_0" bit 10
   5004: 'Carrier 78 Standard Output Card Fault', class No Acknowledgement, trigger "DB302_HMI_Faults_Carrier78_Faults_0" bit 11
   5005: 'Carrier 78 Encoder Position Fault', class No Acknowledgement, trigger "DB302_HMI_Faults_Carrier78_Faults_0" bit 12
   5006: 'Carrier 78 Encoder Internal Error', class No Acknowledgement, trigger "DB302_HMI_Faults_Carrier78_Faults_0" bit 13
   5007: 'Carrier 78 Encoder Comm Fault', class No Acknowledgement, trigger "DB302_HMI_Faults_Carrier78_Faults_0" bit 14
   5008: 'Carrier 78 HMI Comm Fault', class No Acknowledgement, trigger "DB302_HMI_Faults_Carrier78_Faults_0" bit 15
   5009: 'Carrier 78 Crash Detection Fault', class No Acknowledgement, trigger "DB302_HMI_Faults_Carrier78_Faults_1" bit 0
   5010: 'Carrier 78 Carrier Number Invalid', class No Acknowledgement, trigger "DB302_HMI_Faults_Carrier78_Faults_1" bit 1
   5011: 'Carrier 78 Drive: PROFINET configuration error', class No Acknowledgement, trigger "DB302_HMI_Faults_Carrier78_Faults_1" bit 2
   5012: 'Carrier 78 Drive: Error internal communications', class No Acknowledgement, trigger "DB302_HMI_Faults_Carrier78_Faults_1" bit 3
   5013: 'Carrier 78 Drive: Motor overtemperature', class No Acknowledgement, trigger "DB302_HMI_Faults_Carrier78_Faults_1" bit 4
   5014: 'Carrier 78 Drive: Motor overcurrent', class No Acknowledgement, trigger "DB302_HMI_Faults_Carrier78_Faults_1" bit 5
   5015: 'Carrier 78 Drive: Infeed or power unit not ready', class No Acknowledgement, trigger "DB302_HMI_Faults_Carrier78_Faults_1" bit 6
   5016: 'Carrier 78 Drive: Short-circuit/ground fault detected', class No Acknowledgement, trigger "DB302_HMI_Faults_Carrier78_Faults_1" bit 7
   5017: 'Carrier 78 Drive: PROFINET Setpoint timeout', class No Acknowledgement, trigger "DB302_HMI_Faults_Carrier78_Faults_1" bit 8
   5018: 'Carrier 78 Power unit: Overcurrent', class No Acknowledgement, trigger "DB302_HMI_Faults_Carrier78_Faults_1" bit 9
   5019: 'Carrier 78 Power unit: DC link voltage overvoltage', class No Acknowledgement, trigger "DB302_HMI_Faults_Carrier78_Faults_1" bit 10
   5020: 'Carrier 78 Power unit: DC link voltage undervoltage', class No Acknowledgement, trigger "DB302_HMI_Faults_Carrier78_Faults_1" bit 11
   5021: 'Carrier 78 Power unit: Line phase failure in main circuit', class No Acknowledgement, trigger "DB302_HMI_Faults_Carrier78_Faults_1" bit 12
   5022: 'Carrier 78 Power unit: Phase failure motor cable', class No Acknowledgement, trigger "DB302_HMI_Faults_Carrier78_Faults_1" bit 13
   5023: 'Carrier 78 Power unit: Ground fault', class No Acknowledgement, trigger "DB302_HMI_Faults_Carrier78_Faults_1" bit 14
   5024: 'Spare_Fault_5024', class No Acknowledgement, trigger "DB302_HMI_Faults_Carrier78_Faults_1" bit 15
   5025: 'Carrier 78 Motion Off Fault', class No Acknowledgement, trigger "DB302_HMI_Faults_Carrier78_Faults_2" bit 0
   5026: 'Carrier 78 Motion On Fault', class No Acknowledgement, trigger "DB302_HMI_Faults_Carrier78_Faults_2" bit 1
   5027: 'Carrier 78 Spacing Fault', class No Acknowledgement, trigger "DB302_HMI_Faults_Carrier78_Faults_2" bit 2
   5028: 'Carrier 78 Duplicate Carrier Number Fault', class No Acknowledgement, trigger "DB302_HMI_Faults_Carrier78_Faults_2" bit 3
   5029: 'Spare_Fault_5029', class No Acknowledgement, trigger "DB302_HMI_Faults_Carrier78_Faults_2" bit 4
   5030: 'Spare_Fault_5030', class No Acknowledgement, trigger "DB302_HMI_Faults_Carrier78_Faults_2" bit 5
   5031: 'Spare_Fault_5031', class No Acknowledgement, trigger "DB302_HMI_Faults_Carrier78_Faults_2" bit 6
   5032: 'Spare_Fault_5032', class No Acknowledgement, trigger "DB302_HMI_Faults_Carrier78_Faults_2" bit 7
   5033: 'Spare_Fault_5033', class No Acknowledgement, trigger "DB302_HMI_Faults_Carrier78_Faults_2" bit 8
   5034: 'Spare_Fault_5034', class No Acknowledgement, trigger "DB302_HMI_Faults_Carrier78_Faults_2" bit 9
   5035: 'Spare_Fault_5035', class No Acknowledgement, trigger "DB302_HMI_Faults_Carrier78_Faults_2" bit 10
   5036: 'Spare_Fault_5036', class No Acknowledgement, trigger "DB302_HMI_Faults_Carrier78_Faults_2" bit 11
   5037: 'Spare_Fault_5037', class No Acknowledgement, trigger "DB302_HMI_Faults_Carrier78_Faults_2" bit 12
   5038: 'Spare_Fault_5038', class No Acknowledgement, trigger "DB302_HMI_Faults_Carrier78_Faults_2" bit 13
   5039: 'Spare_Fault_5039', class No Acknowledgement, trigger "DB302_HMI_Faults_Carrier78_Faults_2" bit 14
   5040: 'Spare_Fault_5040', class No Acknowledgement, trigger "DB302_HMI_Faults_Carrier78_Faults_2" bit 15
   5041: 'Spare_Fault_5041', class No Acknowledgement, trigger "DB302_HMI_Faults_Carrier78_Faults_3" bit 0
   5042: 'Spare_Fault_5042', class No Acknowledgement, trigger "DB302_HMI_Faults_Carrier78_Faults_3" bit 1
   5043: 'Spare_Fault_5043', class No Acknowledgement, trigger "DB302_HMI_Faults_Carrier78_Faults_3" bit 2
   5044: 'Spare_Fault_5044', class No Acknowledgement, trigger "DB302_HMI_Faults_Carrier78_Faults_3" bit 3
   5045: 'Spare_Fault_5045', class No Acknowledgement, trigger "DB302_HMI_Faults_Carrier78_Faults_3" bit 4
   5046: 'Spare_Fault_5046', class No Acknowledgement, trigger "DB302_HMI_Faults_Carrier78_Faults_3" bit 5
   5047: 'Spare_Fault_5047', class No Acknowledgement, trigger "DB302_HMI_Faults_Carrier78_Faults_3" bit 6
   5048: 'Spare_Fault_5048', class No Acknowledgement, trigger "DB302_HMI_Faults_Carrier78_Faults_3" bit 7
   5049: 'Spare_Fault_5049', class No Acknowledgement, trigger "DB302_HMI_Faults_Carrier78_Faults_3" bit 8
   5050: 'Spare_Fault_5050', class No Acknowledgement, trigger "DB302_HMI_Faults_Carrier78_Faults_3" bit 9
   5051: 'Spare_Fault_5051', class No Acknowledgement, trigger "DB302_HMI_Faults_Carrier78_Faults_3" bit 10
   5052: 'Spare_Fault_5052', class No Acknowledgement, trigger "DB302_HMI_Faults_Carrier78_Faults_3" bit 11
   5053: 'Spare_Fault_5053', class No Acknowledgement, trigger "DB302_HMI_Faults_Carrier78_Faults_3" bit 12
   5054: 'Spare_Fault_5054', class No Acknowledgement, trigger "DB302_HMI_Faults_Carrier78_Faults_3" bit 13
   5055: 'Spare_Fault_5055', class No Acknowledgement, trigger "DB302_HMI_Faults_Carrier78_Faults_3" bit 14
   5056: 'Spare_Fault_5056', class No Acknowledgement, trigger "DB302_HMI_Faults_Carrier78_Faults_3" bit 15
   5057: 'Carrier 79 Disconnect Open Power Fault DI11.0', class No Acknowledgement, trigger "DB302_HMI_Faults_Carrier79_Faults_0" bit 0
   5058: 'Carrier 79 Drive Profinet Comm Fault', class No Acknowledgement, trigger "DB302_HMI_Faults_Carrier79_Faults_0" bit 1
   5059: 'Carrier 79 Production Stop Not Reset', class No Acknowledgement, trigger "DB302_HMI_Faults_Carrier79_Faults_0" bit 2
   5060: 'Carrier 79 CB02122 Tripped', class No Acknowledgement, trigger "DB302_HMI_Faults_Carrier79_Faults_0" bit 3
   5061: 'Carrier 79 CB02123 Tripped', class No Acknowledgement, trigger "DB302_HMI_Faults_Carrier79_Faults_0" bit 4
   5062: 'Carrier 79 AUX1 CB Tripped', class No Acknowledgement, trigger "DB302_HMI_Faults_Carrier79_Faults_0" bit 5
   5063: 'Carrier 79 AUX2 CB Tripped', class No Acknowledgement, trigger "DB302_HMI_Faults_Carrier79_Faults_0" bit 6
   5064: 'Carrier 79 PLC Not Communicating', class No Acknowledgement, trigger "DB302_HMI_Faults_Carrier79_Faults_0" bit 7
   5065: 'Carrier 79 Safe Input Card Fault', class No Acknowledgement, trigger "DB302_HMI_Faults_Carrier79_Faults_0" bit 8
   5066: 'Carrier 79 Safe Output Card Fault', class No Acknowledgement, trigger "DB302_HMI_Faults_Carrier79_Faults_0" bit 9
   5067: 'Carrier 79 Standard Input Card Fault', class No Acknowledgement, trigger "DB302_HMI_Faults_Carrier79_Faults_0" bit 10
   5068: 'Carrier 79 Standard Output Card Fault', class No Acknowledgement, trigger "DB302_HMI_Faults_Carrier79_Faults_0" bit 11
   5069: 'Carrier 79 Encoder Position Fault', class No Acknowledgement, trigger "DB302_HMI_Faults_Carrier79_Faults_0" bit 12
   5070: 'Carrier 79 Encoder Internal Error', class No Acknowledgement, trigger "DB302_HMI_Faults_Carrier79_Faults_0" bit 13
   5071: 'Carrier 79 Encoder Comm Fault', class No Acknowledgement, trigger "DB302_HMI_Faults_Carrier79_Faults_0" bit 14
   5072: 'Carrier 79 HMI Comm Fault', class No Acknowledgement, trigger "DB302_HMI_Faults_Carrier79_Faults_0" bit 15
   5073: 'Carrier 79 Crash Detection Fault', class No Acknowledgement, trigger "DB302_HMI_Faults_Carrier79_Faults_1" bit 0
   5074: 'Carrier 79 Carrier Number Invalid', class No Acknowledgement, trigger "DB302_HMI_Faults_Carrier79_Faults_1" bit 1
   5075: 'Carrier 79 Drive: PROFINET configuration error', class No Acknowledgement, trigger "DB302_HMI_Faults_Carrier79_Faults_1" bit 2
   5076: 'Carrier 79 Drive: Error internal communications', class No Acknowledgement, trigger "DB302_HMI_Faults_Carrier79_Faults_1" bit 3
   5077: 'Carrier 79 Drive: Motor overtemperature', class No Acknowledgement, trigger "DB302_HMI_Faults_Carrier79_Faults_1" bit 4
   5078: 'Carrier 79 Drive: Motor overcurrent', class No Acknowledgement, trigger "DB302_HMI_Faults_Carrier79_Faults_1" bit 5
   5079: 'Carrier 79 Drive: Infeed or power unit not ready', class No Acknowledgement, trigger "DB302_HMI_Faults_Carrier79_Faults_1" bit 6
